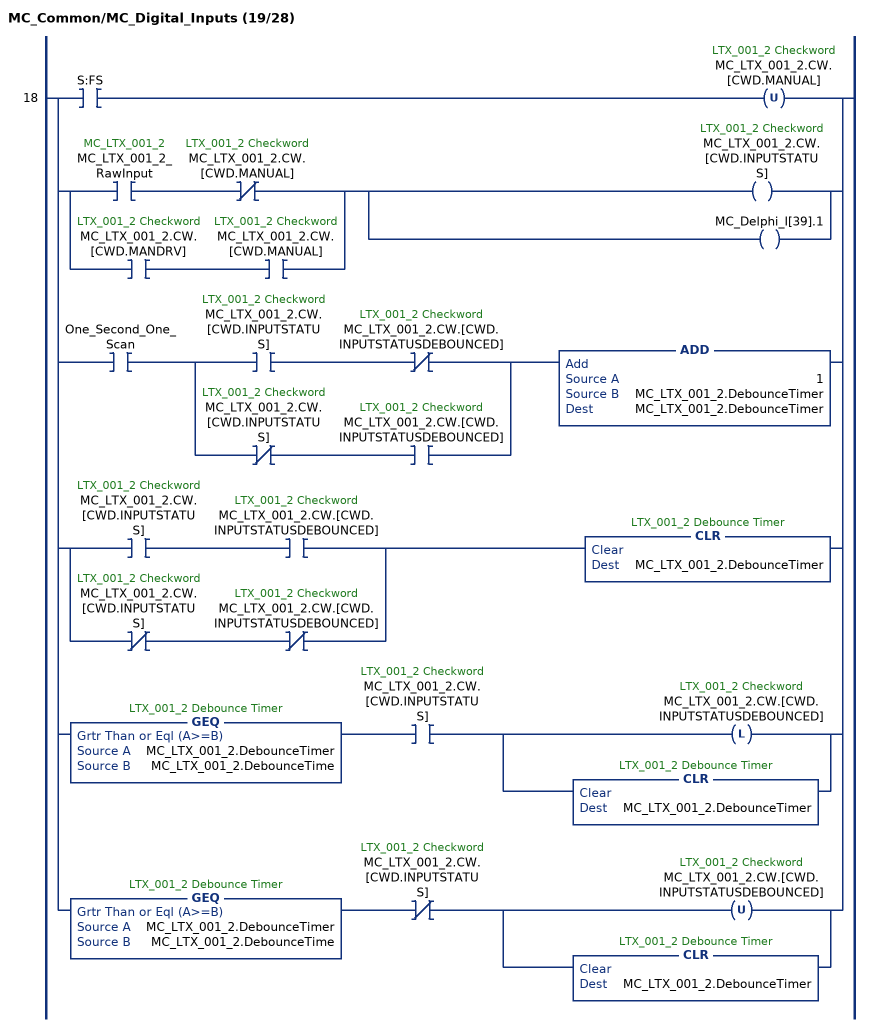
   18: [XIC(S:FS) OTU(MC_LTX_001_2.CW.[CWD.MANUAL]) ,[XIC(MC_LTX_001_2_RawInput) XIO(MC_LTX_001_2.CW.[CWD.MANUAL]) ,XIC(MC_LTX_001_2.CW.[CWD.MANDRV]) XIC(MC_LTX_001_2.CW.[CWD.MANUAL]) ] [OTE(MC_LTX_001_2.CW.[CWD.INPUTSTATUS]) ,OTE(MC_Delphi_I[39].1) ] ,XIC(One_Second_One_Scan) [XIC(MC_LTX_001_2.CW.[CWD.INPUTSTATUS]) XIO(MC_LTX_001_2.CW.[CWD.INPUTSTATUSDEBOUNCED]) ,XIO(MC_LTX_001_2.CW.[CWD.INPUTSTATUS]) XIC(MC_LTX_001_2.CW.[CWD.INPUTSTATUSDEBOUNCED]) ] ADD(1,MC_LTX_001_2.DebounceTimer,MC_LTX_001_2.DebounceTimer) ,[XIC(MC_LTX_001_2.CW.[CWD.INPUTSTATUS]) XIC(MC_LTX_001_2.CW.[CWD.INPUTSTATUSDEBOUNCED]) ,XIO(MC_LTX_001_2.CW.[CWD.INPUTSTATUS]) XIO(MC_LTX_001_2.CW.[CWD.INPUTSTATUSDEBOUNCED]) ] CLR(MC_LTX_001_2.DebounceTimer) ,GEQ(MC_LTX_001_2.DebounceTimer,MC_LTX_001_2.DebounceTime) XIC(MC_LTX_001_2.CW.[CWD.INPUTSTATUS]) [OTL(MC_LTX_001_2.CW.[CWD.INPUTSTATUSDEBOUNCED]) ,CLR(MC_LTX_001_2.DebounceTimer) ] ,GEQ(MC_LTX_001_2.DebounceTimer,MC_LTX_001_2.DebounceTime) XIO(MC_LTX_001_2.CW.[CWD.INPUTSTATUS]) [OTU(MC_LTX_001_2.CW.[CWD.INPUTSTATUSDEBOUNCED]) ,CLR(MC_LTX_001_2.DebounceTimer) ] ];
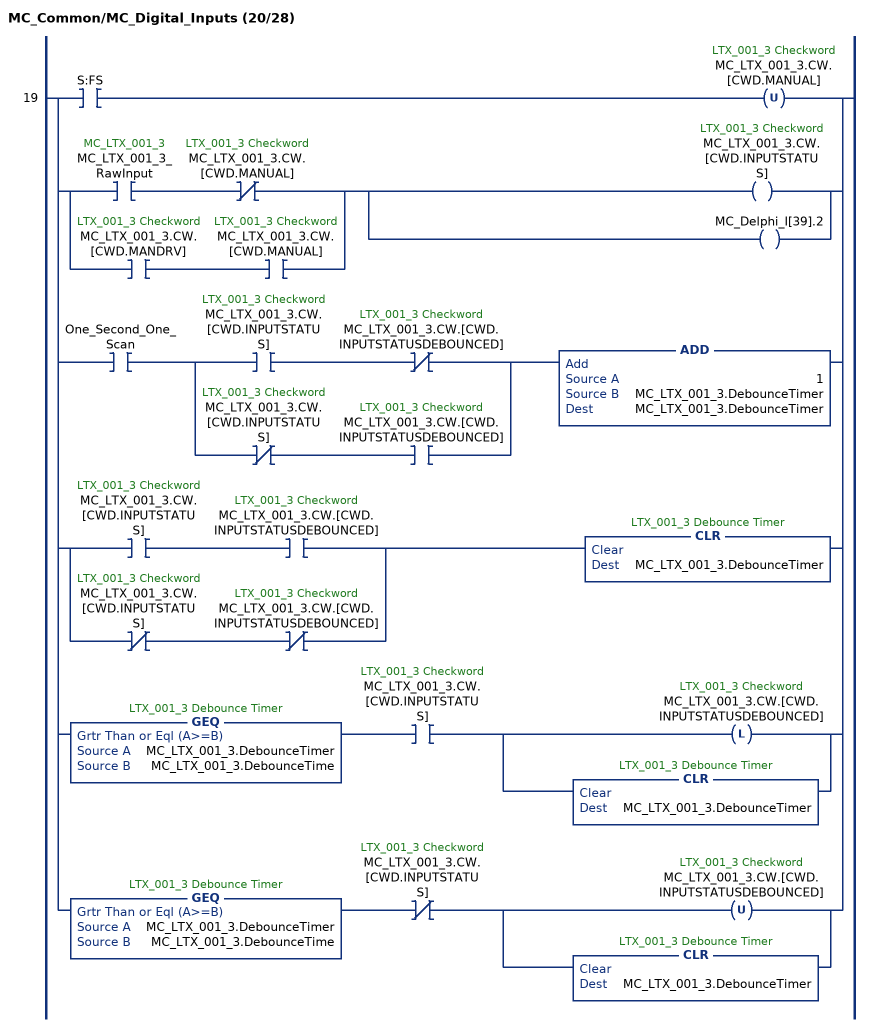
   19: [XIC(S:FS) OTU(MC_LTX_001_3.CW.[CWD.MANUAL]) ,[XIC(MC_LTX_001_3_RawInput) XIO(MC_LTX_001_3.CW.[CWD.MANUAL]) ,XIC(MC_LTX_001_3.CW.[CWD.MANDRV]) XIC(MC_LTX_001_3.CW.[CWD.MANUAL]) ] [OTE(MC_LTX_001_3.CW.[CWD.INPUTSTATUS]) ,OTE(MC_Delphi_I[39].2) ] ,XIC(One_Second_One_Scan) [XIC(MC_LTX_001_3.CW.[CWD.INPUTSTATUS]) XIO(MC_LTX_001_3.CW.[CWD.INPUTSTATUSDEBOUNCED]) ,XIO(MC_LTX_001_3.CW.[CWD.INPUTSTATUS]) XIC(MC_LTX_001_3.CW.[CWD.INPUTSTATUSDEBOUNCED]) ] ADD(1,MC_LTX_001_3.DebounceTimer,MC_LTX_001_3.DebounceTimer) ,[XIC(MC_LTX_001_3.CW.[CWD.INPUTSTATUS]) XIC(MC_LTX_001_3.CW.[CWD.INPUTSTATUSDEBOUNCED]) ,XIO(MC_LTX_001_3.CW.[CWD.INPUTSTATUS]) XIO(MC_LTX_001_3.CW.[CWD.INPUTSTATUSDEBOUNCED]) ] CLR(MC_LTX_001_3.DebounceTimer) ,GEQ(MC_LTX_001_3.DebounceTimer,MC_LTX_001_3.DebounceTime) XIC(MC_LTX_001_3.CW.[CWD.INPUTSTATUS]) [OTL(MC_LTX_001_3.CW.[CWD.INPUTSTATUSDEBOUNCED]) ,CLR(MC_LTX_001_3.DebounceTimer) ] ,GEQ(MC_LTX_001_3.DebounceTimer,MC_LTX_001_3.DebounceTime) XIO(MC_LTX_001_3.CW.[CWD.INPUTSTATUS]) [OTU(MC_LTX_001_3.CW.[CWD.INPUTSTATUSDEBOUNCED]) ,CLR(MC_LTX_001_3.DebounceTimer) ] ];
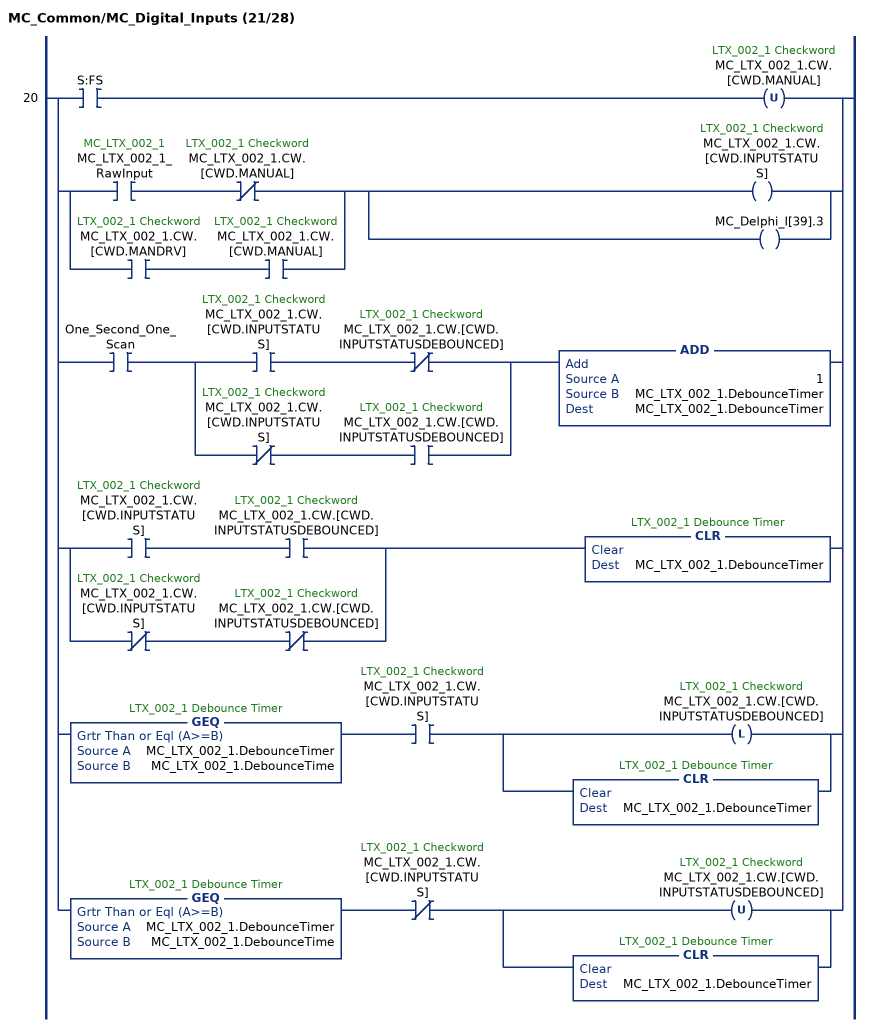
   20: [XIC(S:FS) OTU(MC_LTX_002_1.CW.[CWD.MANUAL]) ,[XIC(MC_LTX_002_1_RawInput) XIO(MC_LTX_002_1.CW.[CWD.MANUAL]) ,XIC(MC_LTX_002_1.CW.[CWD.MANDRV]) XIC(MC_LTX_002_1.CW.[CWD.MANUAL]) ] [OTE(MC_LTX_002_1.CW.[CWD.INPUTSTATUS]) ,OTE(MC_Delphi_I[39].3) ] ,XIC(One_Second_One_Scan) [XIC(MC_LTX_002_1.CW.[CWD.INPUTSTATUS]) XIO(MC_LTX_002_1.CW.[CWD.INPUTSTATUSDEBOUNCED]) ,XIO(MC_LTX_002_1.CW.[CWD.INPUTSTATUS]) XIC(MC_LTX_002_1.CW.[CWD.INPUTSTATUSDEBOUNCED]) ] ADD(1,MC_LTX_002_1.DebounceTimer,MC_LTX_002_1.DebounceTimer) ,[XIC(MC_LTX_002_1.CW.[CWD.INPUTSTATUS]) XIC(MC_LTX_002_1.CW.[CWD.INPUTSTATUSDEBOUNCED]) ,XIO(MC_LTX_002_1.CW.[CWD.INPUTSTATUS]) XIO(MC_LTX_002_1.CW.[CWD.INPUTSTATUSDEBOUNCED]) ] CLR(MC_LTX_002_1.DebounceTimer) ,GEQ(MC_LTX_002_1.DebounceTimer,MC_LTX_002_1.DebounceTime) XIC(MC_LTX_002_1.CW.[CWD.INPUTSTATUS]) [OTL(MC_LTX_002_1.CW.[CWD.INPUTSTATUSDEBOUNCED]) ,CLR(MC_LTX_002_1.DebounceTimer) ] ,GEQ(MC_LTX_002_1.DebounceTimer,MC_LTX_002_1.DebounceTime) XIO(MC_LTX_002_1.CW.[CWD.INPUTSTATUS]) [OTU(MC_LTX_002_1.CW.[CWD.INPUTSTATUSDEBOUNCED]) ,CLR(MC_LTX_002_1.DebounceTimer) ] ];
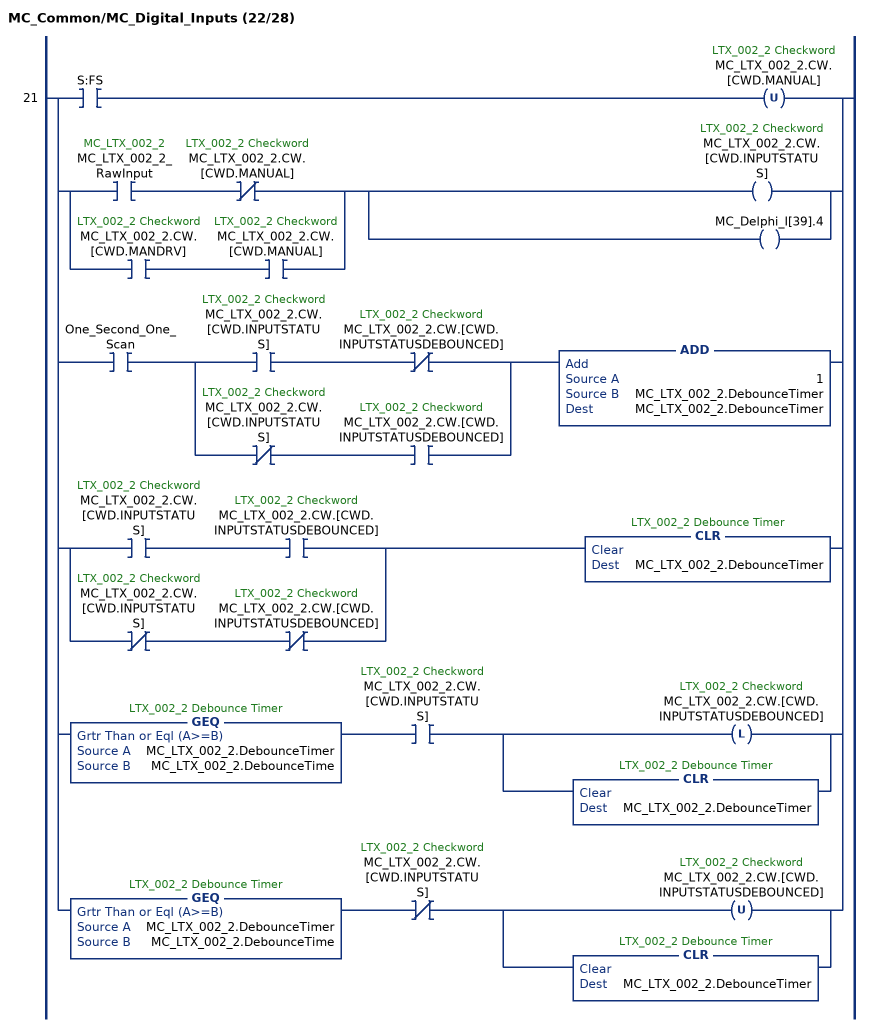
   21: [XIC(S:FS) OTU(MC_LTX_002_2.CW.[CWD.MANUAL]) ,[XIC(MC_LTX_002_2_RawInput) XIO(MC_LTX_002_2.CW.[CWD.MANUAL]) ,XIC(MC_LTX_002_2.CW.[CWD.MANDRV]) XIC(MC_LTX_002_2.CW.[CWD.MANUAL]) ] [OTE(MC_LTX_002_2.CW.[CWD.INPUTSTATUS]) ,OTE(MC_Delphi_I[39].4) ] ,XIC(One_Second_One_Scan) [XIC(MC_LTX_002_2.CW.[CWD.INPUTSTATUS]) XIO(MC_LTX_002_2.CW.[CWD.INPUTSTATUSDEBOUNCED]) ,XIO(MC_LTX_002_2.CW.[CWD.INPUTSTATUS]) XIC(MC_LTX_002_2.CW.[CWD.INPUTSTATUSDEBOUNCED]) ] ADD(1,MC_LTX_002_2.DebounceTimer,MC_LTX_002_2.DebounceTimer) ,[XIC(MC_LTX_002_2.CW.[CWD.INPUTSTATUS]) XIC(MC_LTX_002_2.CW.[CWD.INPUTSTATUSDEBOUNCED]) ,XIO(MC_LTX_002_2.CW.[CWD.INPUTSTATUS]) XIO(MC_LTX_002_2.CW.[CWD.INPUTSTATUSDEBOUNCED]) ] CLR(MC_LTX_002_2.DebounceTimer) ,GEQ(MC_LTX_002_2.DebounceTimer,MC_LTX_002_2.DebounceTime) XIC(MC_LTX_002_2.CW.[CWD.INPUTSTATUS]) [OTL(MC_LTX_002_2.CW.[CWD.INPUTSTATUSDEBOUNCED]) ,CLR(MC_LTX_002_2.DebounceTimer) ] ,GEQ(MC_LTX_002_2.DebounceTimer,MC_LTX_002_2.DebounceTime) XIO(MC_LTX_002_2.CW.[CWD.INPUTSTATUS]) [OTU(MC_LTX_002_2.CW.[CWD.INPUTSTATUSDEBOUNCED]) ,CLR(MC_LTX_002_2.DebounceTimer) ] ];
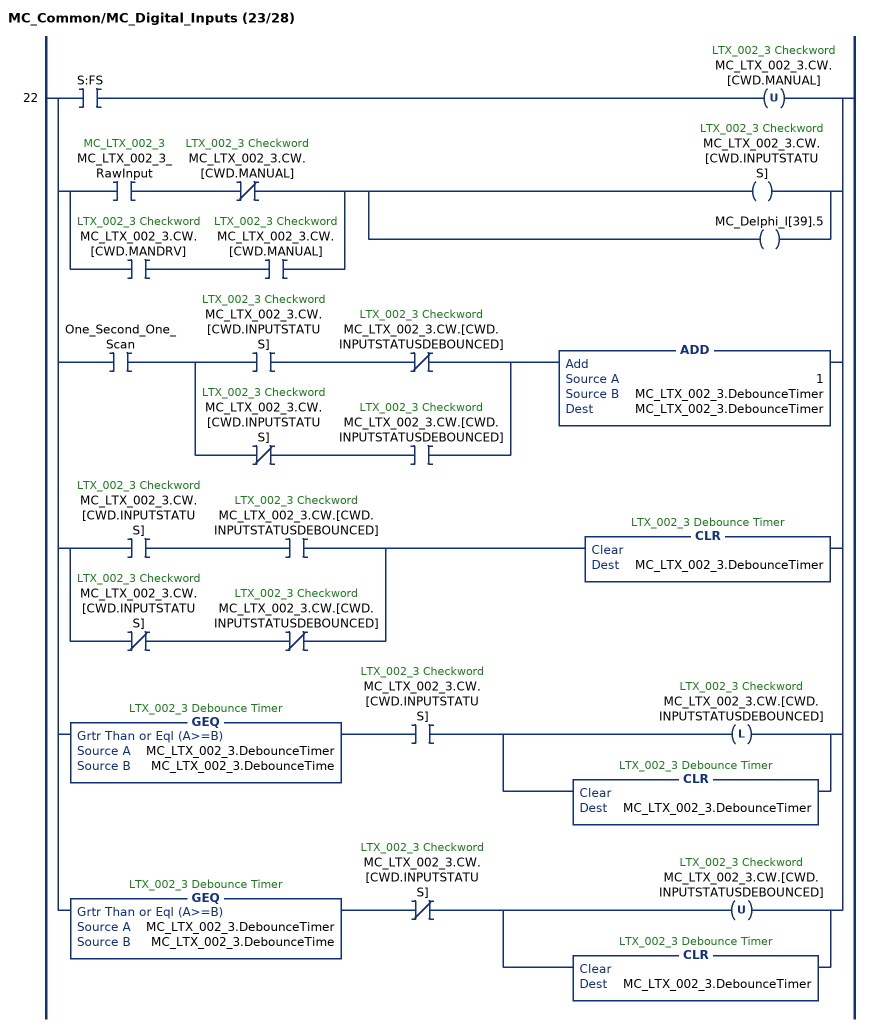
   22: [XIC(S:FS) OTU(MC_LTX_002_3.CW.[CWD.MANUAL]) ,[XIC(MC_LTX_002_3_RawInput) XIO(MC_LTX_002_3.CW.[CWD.MANUAL]) ,XIC(MC_LTX_002_3.CW.[CWD.MANDRV]) XIC(MC_LTX_002_3.CW.[CWD.MANUAL]) ] [OTE(MC_LTX_002_3.CW.[CWD.INPUTSTATUS]) ,OTE(MC_Delphi_I[39].5) ] ,XIC(One_Second_One_Scan) [XIC(MC_LTX_002_3.CW.[CWD.INPUTSTATUS]) XIO(MC_LTX_002_3.CW.[CWD.INPUTSTATUSDEBOUNCED]) ,XIO(MC_LTX_002_3.CW.[CWD.INPUTSTATUS]) XIC(MC_LTX_002_3.CW.[CWD.INPUTSTATUSDEBOUNCED]) ] ADD(1,MC_LTX_002_3.DebounceTimer,MC_LTX_002_3.DebounceTimer) ,[XIC(MC_LTX_002_3.CW.[CWD.INPUTSTATUS]) XIC(MC_LTX_002_3.CW.[CWD.INPUTSTATUSDEBOUNCED]) ,XIO(MC_LTX_002_3.CW.[CWD.INPUTSTATUS]) XIO(MC_LTX_002_3.CW.[CWD.INPUTSTATUSDEBOUNCED]) ] CLR(MC_LTX_002_3.DebounceTimer) ,GEQ(MC_LTX_002_3.DebounceTimer,MC_LTX_002_3.DebounceTime) XIC(MC_LTX_002_3.CW.[CWD.INPUTSTATUS]) [OTL(MC_LTX_002_3.CW.[CWD.INPUTSTATUSDEBOUNCED]) ,CLR(MC_LTX_002_3.DebounceTimer) ] ,GEQ(MC_LTX_002_3.DebounceTimer,MC_LTX_002_3.DebounceTime) XIO(MC_LTX_002_3.CW.[CWD.INPUTSTATUS]) [OTU(MC_LTX_002_3.CW.[CWD.INPUTSTATUSDEBOUNCED]) ,CLR(MC_LTX_002_3.DebounceTimer) ] ];
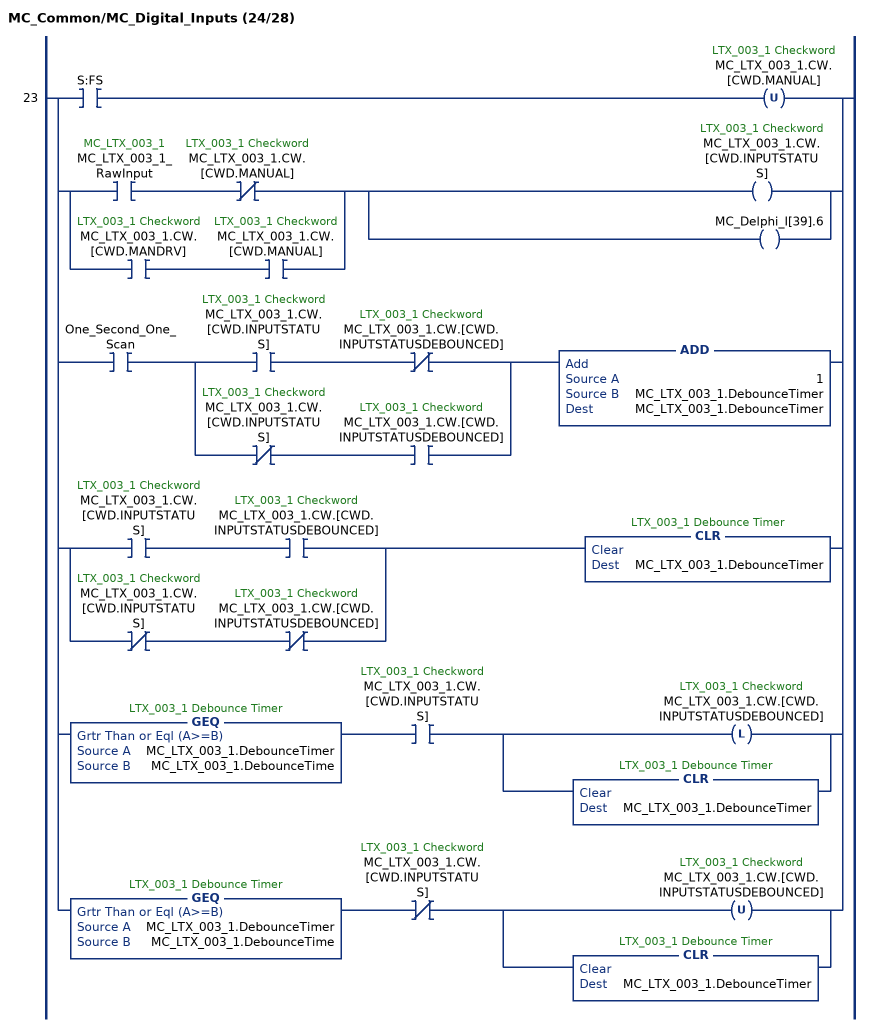
   23: [XIC(S:FS) OTU(MC_LTX_003_1.CW.[CWD.MANUAL]) ,[XIC(MC_LTX_003_1_RawInput) XIO(MC_LTX_003_1.CW.[CWD.MANUAL]) ,XIC(MC_LTX_003_1.CW.[CWD.MANDRV]) XIC(MC_LTX_003_1.CW.[CWD.MANUAL]) ] [OTE(MC_LTX_003_1.CW.[CWD.INPUTSTATUS]) ,OTE(MC_Delphi_I[39].6) ] ,XIC(One_Second_One_Scan) [XIC(MC_LTX_003_1.CW.[CWD.INPUTSTATUS]) XIO(MC_LTX_003_1.CW.[CWD.INPUTSTATUSDEBOUNCED]) ,XIO(MC_LTX_003_1.CW.[CWD.INPUTSTATUS]) XIC(MC_LTX_003_1.CW.[CWD.INPUTSTATUSDEBOUNCED]) ] ADD(1,MC_LTX_003_1.DebounceTimer,MC_LTX_003_1.DebounceTimer) ,[XIC(MC_LTX_003_1.CW.[CWD.INPUTSTATUS]) XIC(MC_LTX_003_1.CW.[CWD.INPUTSTATUSDEBOUNCED]) ,XIO(MC_LTX_003_1.CW.[CWD.INPUTSTATUS]) XIO(MC_LTX_003_1.CW.[CWD.INPUTSTATUSDEBOUNCED]) ] CLR(MC_LTX_003_1.DebounceTimer) ,GEQ(MC_LTX_003_1.DebounceTimer,MC_LTX_003_1.DebounceTime) XIC(MC_LTX_003_1.CW.[CWD.INPUTSTATUS]) [OTL(MC_LTX_003_1.CW.[CWD.INPUTSTATUSDEBOUNCED]) ,CLR(MC_LTX_003_1.DebounceTimer) ] ,GEQ(MC_LTX_003_1.DebounceTimer,MC_LTX_003_1.DebounceTime) XIO(MC_LTX_003_1.CW.[CWD.INPUTSTATUS]) [OTU(MC_LTX_003_1.CW.[CWD.INPUTSTATUSDEBOUNCED]) ,CLR(MC_LTX_003_1.DebounceTimer) ] ];
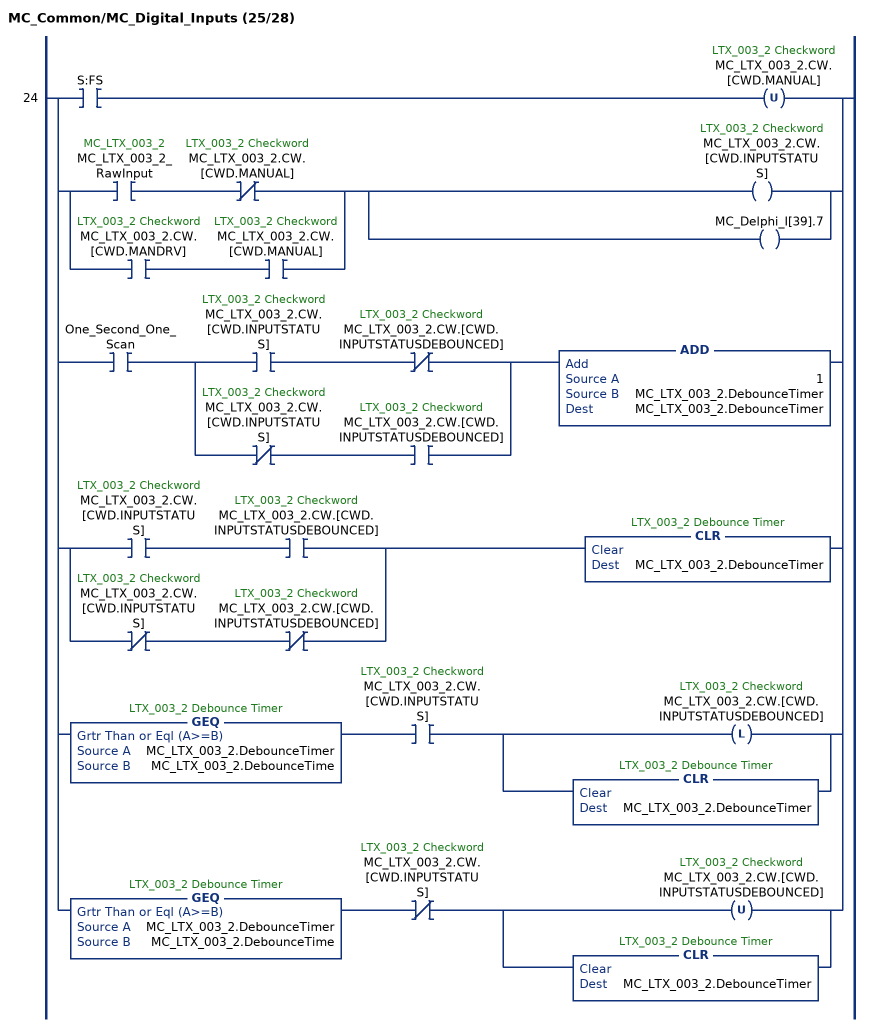
   24: [XIC(S:FS) OTU(MC_LTX_003_2.CW.[CWD.MANUAL]) ,[XIC(MC_LTX_003_2_RawInput) XIO(MC_LTX_003_2.CW.[CWD.MANUAL]) ,XIC(MC_LTX_003_2.CW.[CWD.MANDRV]) XIC(MC_LTX_003_2.CW.[CWD.MANUAL]) ] [OTE(MC_LTX_003_2.CW.[CWD.INPUTSTATUS]) ,OTE(MC_Delphi_I[39].7) ] ,XIC(One_Second_One_Scan) [XIC(MC_LTX_003_2.CW.[CWD.INPUTSTATUS]) XIO(MC_LTX_003_2.CW.[CWD.INPUTSTATUSDEBOUNCED]) ,XIO(MC_LTX_003_2.CW.[CWD.INPUTSTATUS]) XIC(MC_LTX_003_2.CW.[CWD.INPUTSTATUSDEBOUNCED]) ] ADD(1,MC_LTX_003_2.DebounceTimer,MC_LTX_003_2.DebounceTimer) ,[XIC(MC_LTX_003_2.CW.[CWD.INPUTSTATUS]) XIC(MC_LTX_003_2.CW.[CWD.INPUTSTATUSDEBOUNCED]) ,XIO(MC_LTX_003_2.CW.[CWD.INPUTSTATUS]) XIO(MC_LTX_003_2.CW.[CWD.INPUTSTATUSDEBOUNCED]) ] CLR(MC_LTX_003_2.DebounceTimer) ,GEQ(MC_LTX_003_2.DebounceTimer,MC_LTX_003_2.DebounceTime) XIC(MC_LTX_003_2.CW.[CWD.INPUTSTATUS]) [OTL(MC_LTX_003_2.CW.[CWD.INPUTSTATUSDEBOUNCED]) ,CLR(MC_LTX_003_2.DebounceTimer) ] ,GEQ(MC_LTX_003_2.DebounceTimer,MC_LTX_003_2.DebounceTime) XIO(MC_LTX_003_2.CW.[CWD.INPUTSTATUS]) [OTU(MC_LTX_003_2.CW.[CWD.INPUTSTATUSDEBOUNCED]) ,CLR(MC_LTX_003_2.DebounceTimer) ] ];
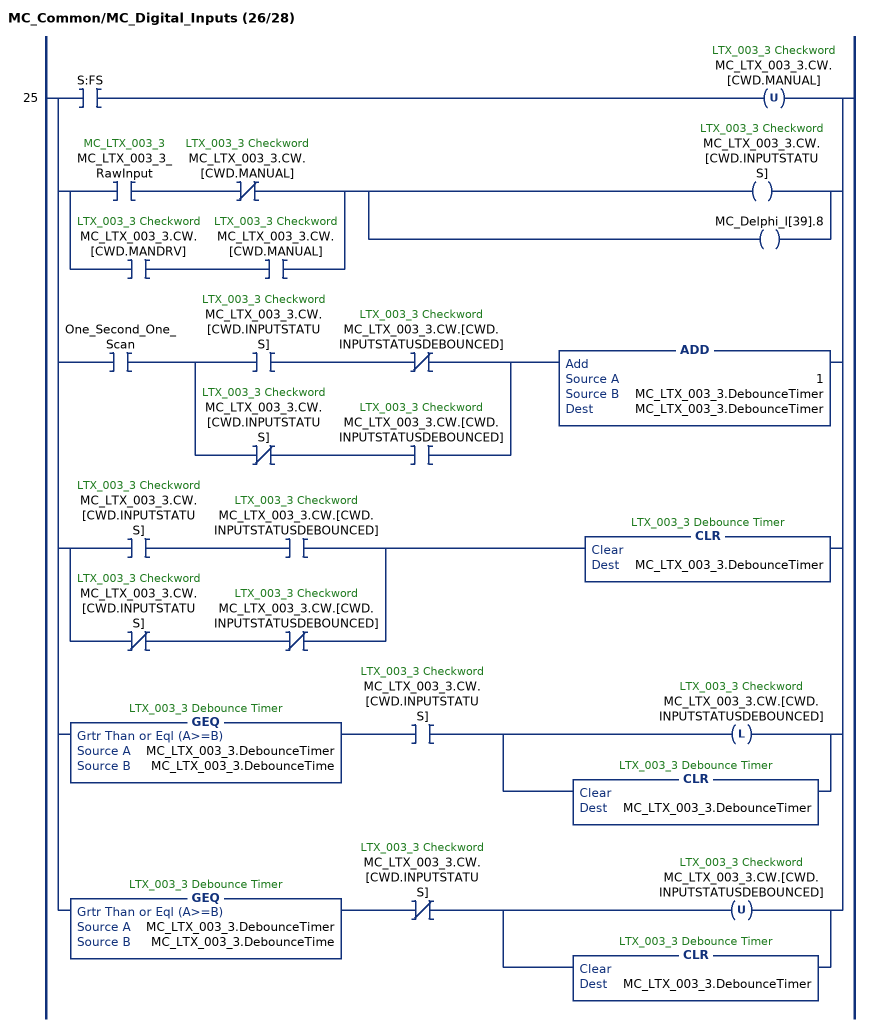
   25: [XIC(S:FS) OTU(MC_LTX_003_3.CW.[CWD.MANUAL]) ,[XIC(MC_LTX_003_3_RawInput) XIO(MC_LTX_003_3.CW.[CWD.MANUAL]) ,XIC(MC_LTX_003_3.CW.[CWD.MANDRV]) XIC(MC_LTX_003_3.CW.[CWD.MANUAL]) ] [OTE(MC_LTX_003_3.CW.[CWD.INPUTSTATUS]) ,OTE(MC_Delphi_I[39].8) ] ,XIC(One_Second_One_Scan) [XIC(MC_LTX_003_3.CW.[CWD.INPUTSTATUS]) XIO(MC_LTX_003_3.CW.[CWD.INPUTSTATUSDEBOUNCED]) ,XIO(MC_LTX_003_3.CW.[CWD.INPUTSTATUS]) XIC(MC_LTX_003_3.CW.[CWD.INPUTSTATUSDEBOUNCED]) ] ADD(1,MC_LTX_003_3.DebounceTimer,MC_LTX_003_3.DebounceTimer) ,[XIC(MC_LTX_003_3.CW.[CWD.INPUTSTATUS]) XIC(MC_LTX_003_3.CW.[CWD.INPUTSTATUSDEBOUNCED]) ,XIO(MC_LTX_003_3.CW.[CWD.INPUTSTATUS]) XIO(MC_LTX_003_3.CW.[CWD.INPUTSTATUSDEBOUNCED]) ] CLR(MC_LTX_003_3.DebounceTimer) ,GEQ(MC_LTX_003_3.DebounceTimer,MC_LTX_003_3.DebounceTime) XIC(MC_LTX_003_3.CW.[CWD.INPUTSTATUS]) [OTL(MC_LTX_003_3.CW.[CWD.INPUTSTATUSDEBOUNCED]) ,CLR(MC_LTX_003_3.DebounceTimer) ] ,GEQ(MC_LTX_003_3.DebounceTimer,MC_LTX_003_3.DebounceTime) XIO(MC_LTX_003_3.CW.[CWD.INPUTSTATUS]) [OTU(MC_LTX_003_3.CW.[CWD.INPUTSTATUSDEBOUNCED]) ,CLR(MC_LTX_003_3.DebounceTimer) ] ];
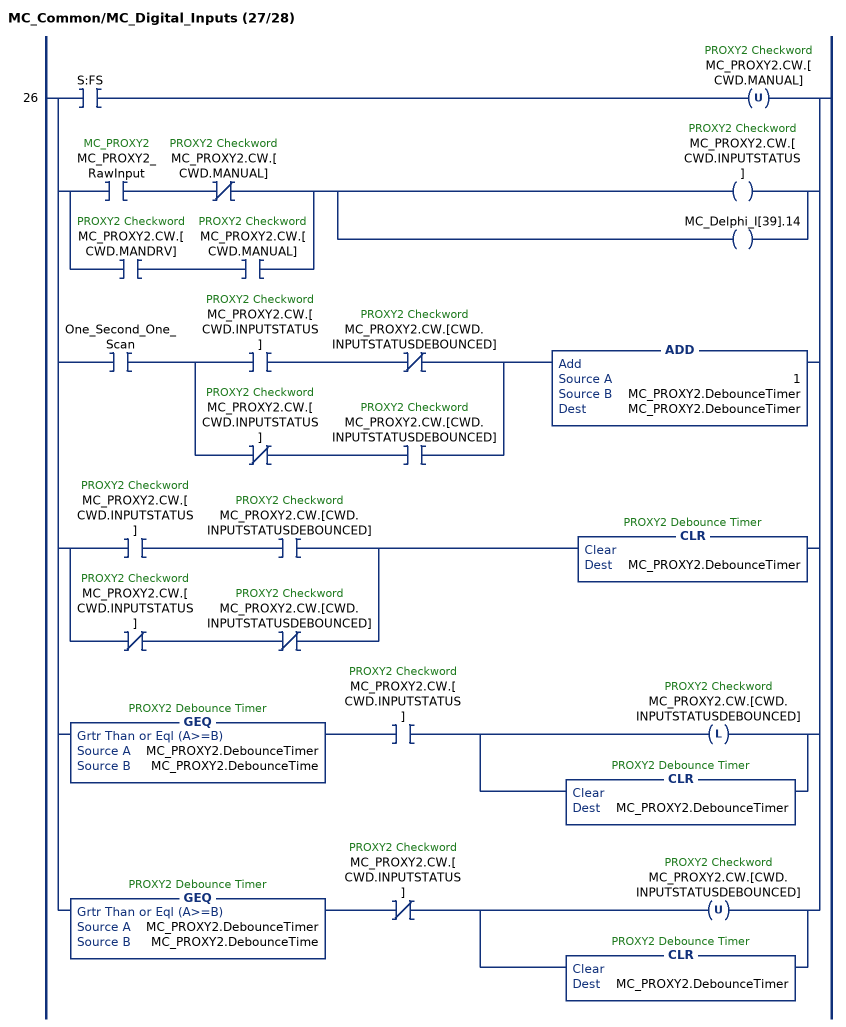
   26: [XIC(S:FS) OTU(MC_PROXY2.CW.[CWD.MANUAL]) ,[XIC(MC_PROXY2_RawInput) XIO(MC_PROXY2.CW.[CWD.MANUAL]) ,XIC(MC_PROXY2.CW.[CWD.MANDRV]) XIC(MC_PROXY2.CW.[CWD.MANUAL]) ] [OTE(MC_PROXY2.CW.[CWD.INPUTSTATUS]) ,OTE(MC_Delphi_I[39].14) ] ,XIC(One_Second_One_Scan) [XIC(MC_PROXY2.CW.[CWD.INPUTSTATUS]) XIO(MC_PROXY2.CW.[CWD.INPUTSTATUSDEBOUNCED]) ,XIO(MC_PROXY2.CW.[CWD.INPUTSTATUS]) XIC(MC_PROXY2.CW.[CWD.INPUTSTATUSDEBOUNCED]) ] ADD(1,MC_PROXY2.DebounceTimer,MC_PROXY2.DebounceTimer) ,[XIC(MC_PROXY2.CW.[CWD.INPUTSTATUS]) XIC(MC_PROXY2.CW.[CWD.INPUTSTATUSDEBOUNCED]) ,XIO(MC_PROXY2.CW.[CWD.INPUTSTATUS]) XIO(MC_PROXY2.CW.[CWD.INPUTSTATUSDEBOUNCED]) ] CLR(MC_PROXY2.DebounceTimer) ,GEQ(MC_PROXY2.DebounceTimer,MC_PROXY2.DebounceTime) XIC(MC_PROXY2.CW.[CWD.INPUTSTATUS]) [OTL(MC_PROXY2.CW.[CWD.INPUTSTATUSDEBOUNCED]) ,CLR(MC_PROXY2.DebounceTimer) ] ,GEQ(MC_PROXY2.DebounceTimer,MC_PROXY2.DebounceTime) XIO(MC_PROXY2.CW.[CWD.INPUTSTATUS]) [OTU(MC_PROXY2.CW.[CWD.INPUTSTATUSDEBOUNCED]) ,CLR(MC_PROXY2.DebounceTimer) ] ];
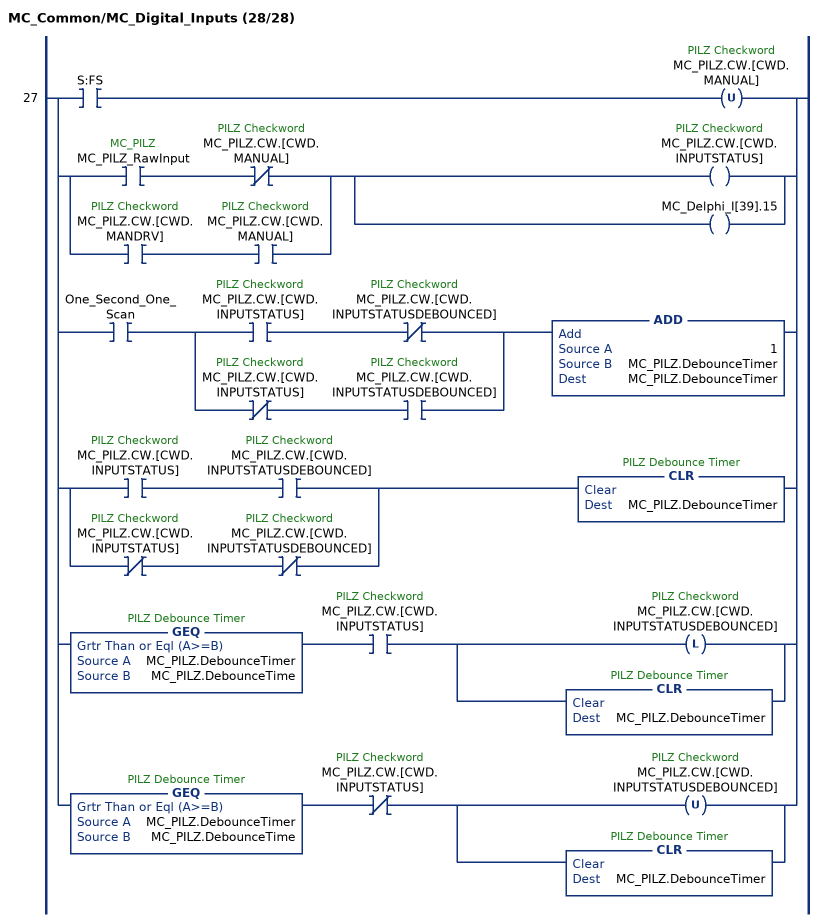
   27: [XIC(S:FS) OTU(MC_PILZ.CW.[CWD.MANUAL]) ,[XIC(MC_PILZ_RawInput) XIO(MC_PILZ.CW.[CWD.MANUAL]) ,XIC(MC_PILZ.CW.[CWD.MANDRV]) XIC(MC_PILZ.CW.[CWD.MANUAL]) ] [OTE(MC_PILZ.CW.[CWD.INPUTSTATUS]) ,OTE(MC_Delphi_I[39].15) ] ,XIC(One_Second_One_Scan) [XIC(MC_PILZ.CW.[CWD.INPUTSTATUS]) XIO(MC_PILZ.CW.[CWD.INPUTSTATUSDEBOUNCED]) ,XIO(MC_PILZ.CW.[CWD.INPUTSTATUS]) XIC(MC_PILZ.CW.[CWD.INPUTSTATUSDEBOUNCED]) ] ADD(1,MC_PILZ.DebounceTimer,MC_PILZ.DebounceTimer) ,[XIC(MC_PILZ.CW.[CWD.INPUTSTATUS]) XIC(MC_PILZ.CW.[CWD.INPUTSTATUSDEBOUNCED]) ,XIO(MC_PILZ.CW.[CWD.INPUTSTATUS]) XIO(MC_PILZ.CW.[CWD.INPUTSTATUSDEBOUNCED]) ] CLR(MC_PILZ.DebounceTimer) ,GEQ(MC_PILZ.DebounceTimer,MC_PILZ.DebounceTime) XIC(MC_PILZ.CW.[CWD.INPUTSTATUS]) [OTL(MC_PILZ.CW.[CWD.INPUTSTATUSDEBOUNCED]) ,CLR(MC_PILZ.DebounceTimer) ] ,GEQ(MC_PILZ.DebounceTimer,MC_PILZ.DebounceTime) XIO(MC_PILZ.CW.[CWD.INPUTSTATUS]) [OTU(MC_PILZ.CW.[CWD.INPUTSTATUSDEBOUNCED]) ,CLR(MC_PILZ.DebounceTimer) ] ];
END_ROUTINE
